(* Logix 5000 project; controller MV vendor 1 type 14 code 217 rev 31.11; software revision 31.00; part 17 of 53 *)
(* tags used below, declared in another part *)
   Alarm_Reset : BOOL;
   CheckTimeMask : INT;
   CLOCKsetvalues : DINT[7];
   CurrentTime : DateTime;
   CWD : CHECKWORD_FLAGS;
   Delphi_Does_Eng_Func : BOOL;
   MC_CLOCK_system_set : BOOL;
   MC_CP1 : PlantItem;   // CP1
   MC_data_file_value_to_move : DINT;
   MC_GBYV1 : PlantItem;   // GBYV1
   MC_N10 : INT[255];   // SETTINGS
   MC_N200 : INT[255];   // CHK_WORK Plant item fault che cking work area
   MC_N255 : INT[255];   // CHECKWORDS Plant item checkword s
   MC_P1 : PlantItem;   // P1
   MC_P2 : PlantItem;   // P2
   MC_P3 : PlantItem;   // P3
   MC_P4 : PlantItem;   // P4
   MC_SFile : INT[255];   // SLC Equivalent System File, So Original Code Can Remain
   MC_SP_R1_1 : PlantItem;   // SP_R1_1
   MC_SP_R2_1 : PlantItem;   // SP_R2_1
   MC_SP_R3_1 : PlantItem;   // SP_R3_1
   MC_T4 : TIMER[255];   // TIMER
   TempChecktime : DINT;
(* MC_Common, continued *)

ROUTINE MC_ITEMCHECK_200   (* ladder *)
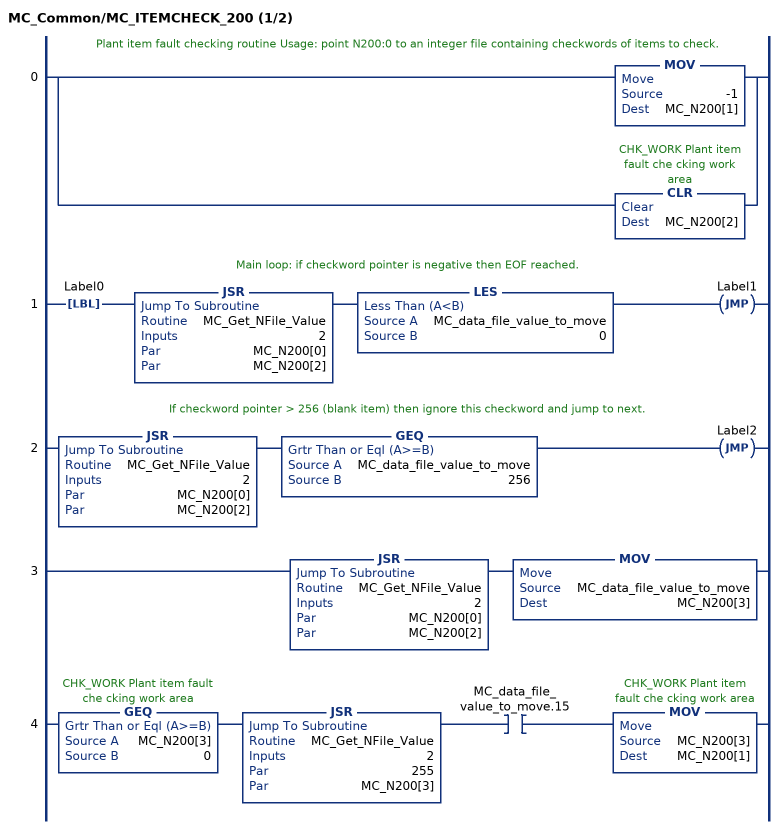
   // Plant item fault checking routine Usage: point N200:0 to an integer file containing checkwords of items to check.
   0: [MOV(-1,MC_N200[1]) ,CLR(MC_N200[2]) ];
   // Main loop: if checkword pointer is negative then EOF reached.
   1: LBL(Label0)JSR(MC_Get_NFile_Value,2,MC_N200[0],MC_N200[2])LES(MC_data_file_value_to_move,0)JMP(Label1);
   // If checkword pointer > 256 (blank item) then ignore this checkword and jump to next.
   2: JSR(MC_Get_NFile_Value,2,MC_N200[0],MC_N200[2])GEQ(MC_data_file_value_to_move,256)JMP(Label2);
   3: JSR(MC_Get_NFile_Value,2,MC_N200[0],MC_N200[2])MOV(MC_data_file_value_to_move,MC_N200[3]);
   4: GEQ(MC_N200[3],0)JSR(MC_Get_NFile_Value,2,255,MC_N200[3])XIC(MC_data_file_value_to_move.15)MOV(MC_N200[3],MC_N200[1]);
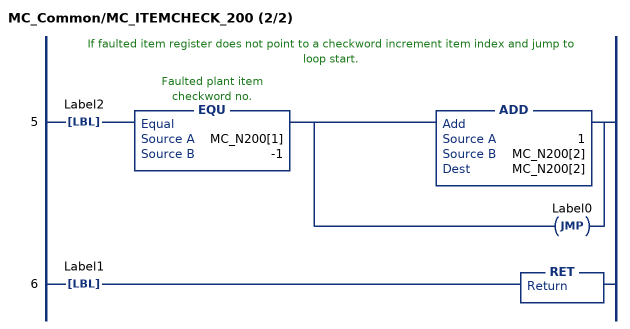
   // If faulted item register does not point to a checkword increment item index and jump to loop start.
   5: LBL(Label2)EQU(MC_N200[1],-1)[ADD(1,MC_N200[2],MC_N200[2]) ,JMP(Label0) ];
   6: LBL(Label1)RET();
END_ROUTINE

ROUTINE MC_MAIN   (* ladder *)
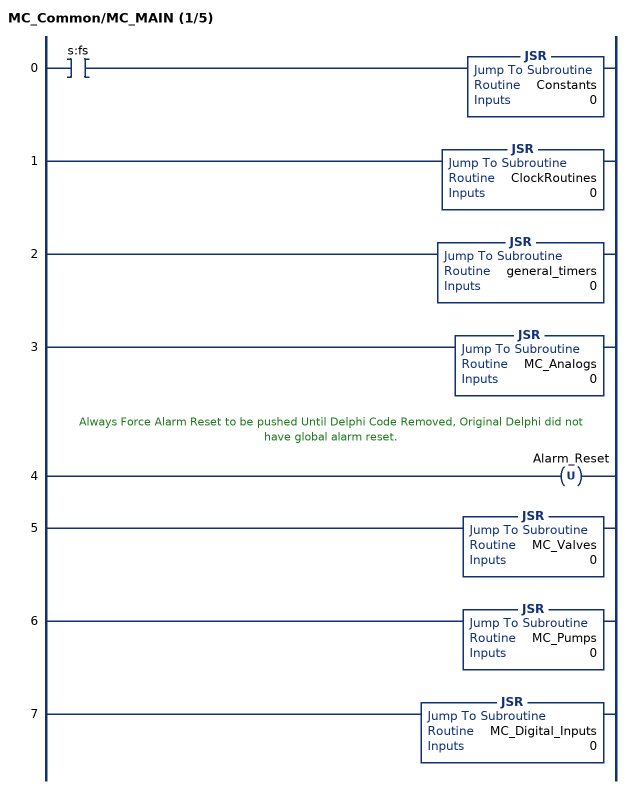
   0: XIC(s:fs)JSR(Constants,0);
   1: JSR(ClockRoutines,0);
   2: JSR(general_timers,0);
   3: JSR(MC_Analogs,0);
   // Always Force Alarm Reset to be pushed Until Delphi Code Removed, Original Delphi did not have global alarm reset.
   4: OTU(Alarm_Reset);
   5: JSR(MC_Valves,0);
   6: JSR(MC_Pumps,0);
   7: JSR(MC_Digital_Inputs,0);
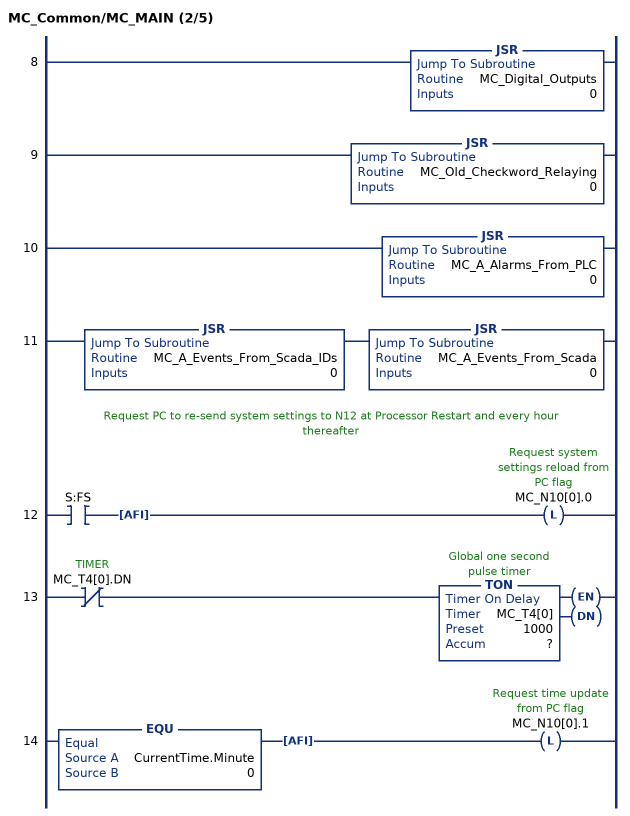
   8: JSR(MC_Digital_Outputs,0);
   9: JSR(MC_Old_Checkword_Relaying,0);
   10: JSR(MC_A_Alarms_From_PLC,0);
   11: JSR(MC_A_Events_From_Scada_IDs,0)JSR(MC_A_Events_From_Scada,0);
   // Request PC to re-send system settings to N12 at Processor Restart and every hour thereafter
   12: XIC(S:FS)AFI()OTL(MC_N10[0].0);
   13: XIO(MC_T4[0].DN)TON(MC_T4[0],?,?);
   14: EQU(CurrentTime.Minute,0)AFI()OTL(MC_N10[0].1);
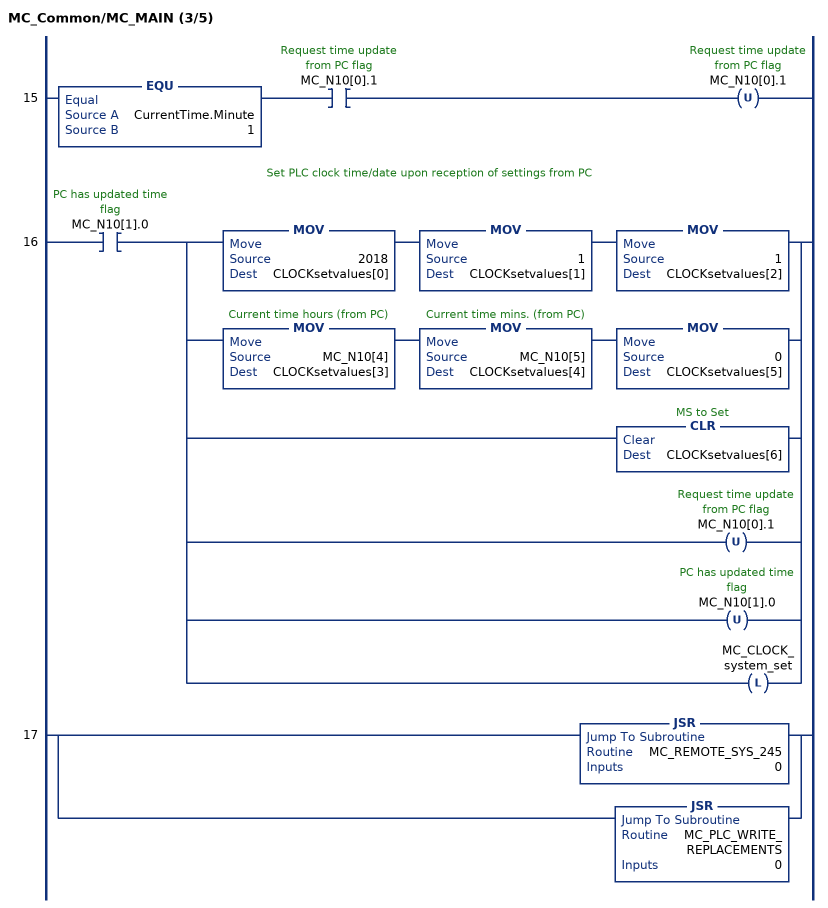
   15: EQU(CurrentTime.Minute,1)XIC(MC_N10[0].1)OTU(MC_N10[0].1);
   // Set PLC clock time/date upon reception of settings from PC
   16: XIC(MC_N10[1].0)[MOV(2018,CLOCKsetvalues[0]) MOV(1,CLOCKsetvalues[1]) MOV(1,CLOCKsetvalues[2]) ,MOV(MC_N10[4],CLOCKsetvalues[3]) MOV(MC_N10[5],CLOCKsetvalues[4]) MOV(0,CLOCKsetvalues[5]) ,CLR(CLOCKsetvalues[6]) ,OTU(MC_N10[0].1) ,OTU(MC_N10[1].0) ,OTL(MC_CLOCK_system_set) ];
   17: [JSR(MC_REMOTE_SYS_245,0) ,JSR(MC_PLC_WRITE_REPLACEMENTS,0) ];
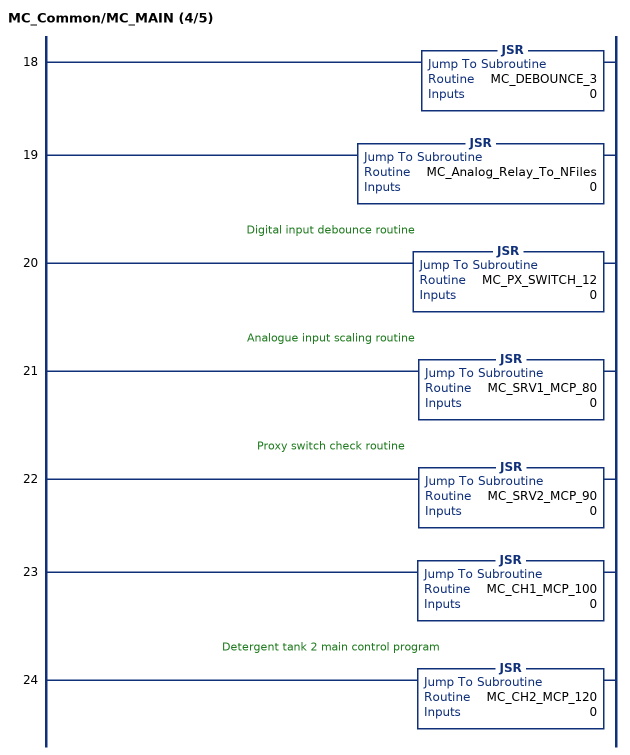
   18: JSR(MC_DEBOUNCE_3,0);
   19: JSR(MC_Analog_Relay_To_NFiles,0);
   // Digital input debounce routine
   20: JSR(MC_PX_SWITCH_12,0);
   // Analogue input scaling routine
   21: JSR(MC_SRV1_MCP_80,0);
   // Proxy switch check routine
   22: JSR(MC_SRV2_MCP_90,0);
   23: JSR(MC_CH1_MCP_100,0);
   // Detergent tank 2 main control program
   24: JSR(MC_CH2_MCP_120,0);
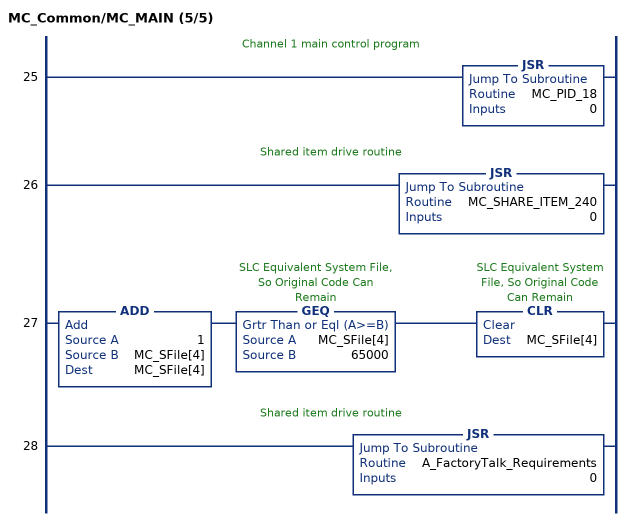
   // Channel 1 main control program
   25: JSR(MC_PID_18,0);
   // Shared item drive routine
   26: JSR(MC_SHARE_ITEM_240,0);
   27: ADD(1,MC_SFile[4],MC_SFile[4])GEQ(MC_SFile[4],65000)CLR(MC_SFile[4]);
   // Shared item drive routine
   28: JSR(A_FactoryTalk_Requirements,0);
END_ROUTINE

ROUTINE MC_Old_Checkword_Relaying   (* ladder *)
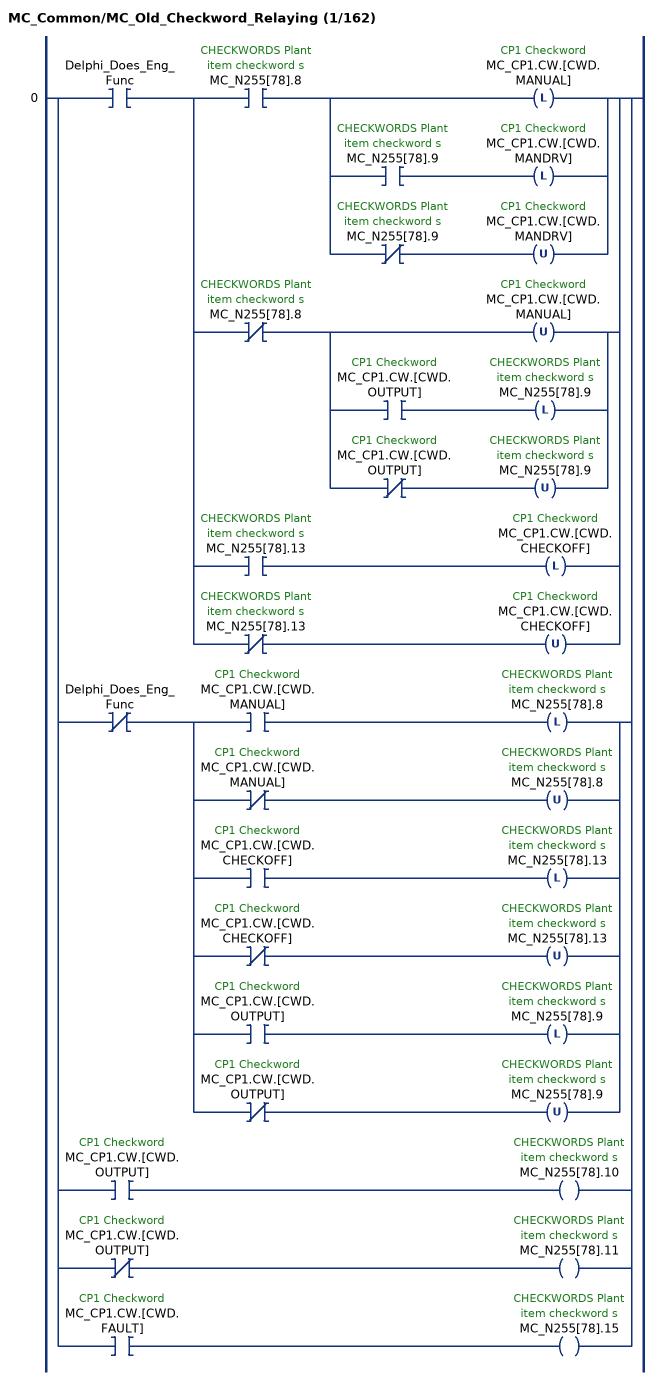
   0: [XIC(Delphi_Does_Eng_Func) [[XIC(MC_N255[78].8) [OTL(MC_CP1.CW.[CWD.MANUAL]) ,XIC(MC_N255[78].9) OTL(MC_CP1.CW.[CWD.MANDRV]) ,XIO(MC_N255[78].9) OTU(MC_CP1.CW.[CWD.MANDRV]) ] ,XIO(MC_N255[78].8) [OTU(MC_CP1.CW.[CWD.MANUAL]) ,[XIC(MC_CP1.CW.[CWD.OUTPUT]) OTL(MC_N255[78].9) ,XIO(MC_CP1.CW.[CWD.OUTPUT]) OTU(MC_N255[78].9) ] ] ] ,[XIC(MC_N255[78].13) OTL(MC_CP1.CW.[CWD.CHECKOFF]) ,XIO(MC_N255[78].13) OTU(MC_CP1.CW.[CWD.CHECKOFF]) ] ] ,XIO(Delphi_Does_Eng_Func) [[XIC(MC_CP1.CW.[CWD.MANUAL]) OTL(MC_N255[78].8) ,XIO(MC_CP1.CW.[CWD.MANUAL]) OTU(MC_N255[78].8) ] ,[XIC(MC_CP1.CW.[CWD.CHECKOFF]) OTL(MC_N255[78].13) ,XIO(MC_CP1.CW.[CWD.CHECKOFF]) OTU(MC_N255[78].13) ] ,[XIC(MC_CP1.CW.[CWD.OUTPUT]) OTL(MC_N255[78].9) ,XIO(MC_CP1.CW.[CWD.OUTPUT]) OTU(MC_N255[78].9) ] ] ,XIC(MC_CP1.CW.[CWD.OUTPUT]) OTE(MC_N255[78].10) ,XIO(MC_CP1.CW.[CWD.OUTPUT]) OTE(MC_N255[78].11) ,XIC(MC_CP1.CW.[CWD.FAULT]) OTE(MC_N255[78].15) ];
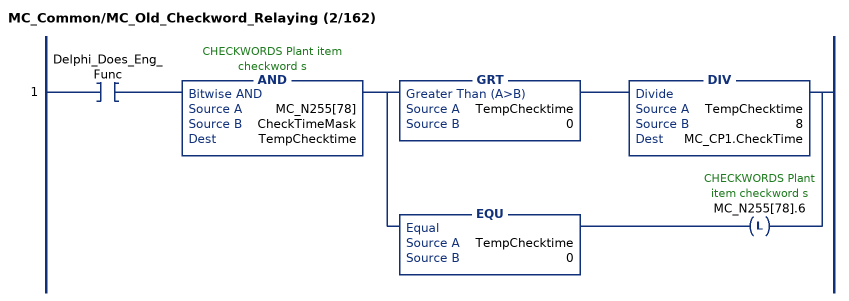
   1: XIC(Delphi_Does_Eng_Func)AND(MC_N255[78],CheckTimeMask,TempChecktime)[GRT(TempChecktime,0) DIV(TempChecktime,8,MC_CP1.CheckTime) ,EQU(TempChecktime,0) OTL(MC_N255[78].6) ];
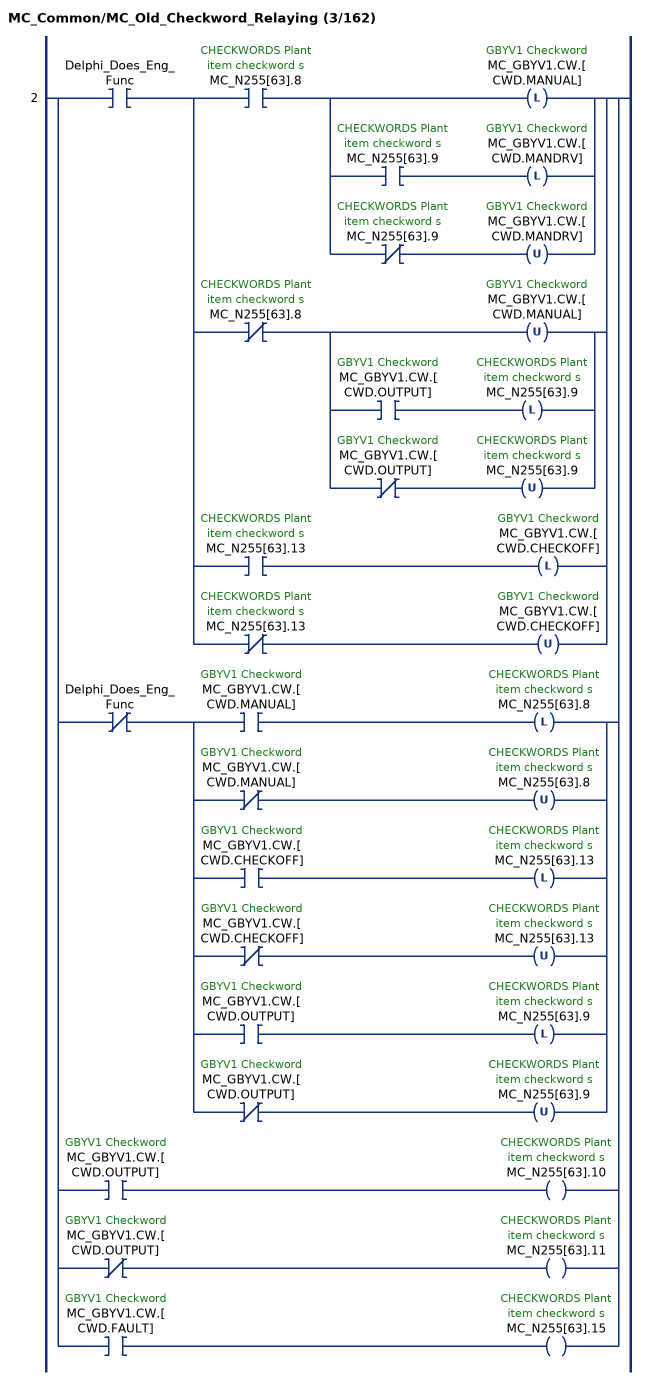
   2: [XIC(Delphi_Does_Eng_Func) [[XIC(MC_N255[63].8) [OTL(MC_GBYV1.CW.[CWD.MANUAL]) ,XIC(MC_N255[63].9) OTL(MC_GBYV1.CW.[CWD.MANDRV]) ,XIO(MC_N255[63].9) OTU(MC_GBYV1.CW.[CWD.MANDRV]) ] ,XIO(MC_N255[63].8) [OTU(MC_GBYV1.CW.[CWD.MANUAL]) ,[XIC(MC_GBYV1.CW.[CWD.OUTPUT]) OTL(MC_N255[63].9) ,XIO(MC_GBYV1.CW.[CWD.OUTPUT]) OTU(MC_N255[63].9) ] ] ] ,[XIC(MC_N255[63].13) OTL(MC_GBYV1.CW.[CWD.CHECKOFF]) ,XIO(MC_N255[63].13) OTU(MC_GBYV1.CW.[CWD.CHECKOFF]) ] ] ,XIO(Delphi_Does_Eng_Func) [[XIC(MC_GBYV1.CW.[CWD.MANUAL]) OTL(MC_N255[63].8) ,XIO(MC_GBYV1.CW.[CWD.MANUAL]) OTU(MC_N255[63].8) ] ,[XIC(MC_GBYV1.CW.[CWD.CHECKOFF]) OTL(MC_N255[63].13) ,XIO(MC_GBYV1.CW.[CWD.CHECKOFF]) OTU(MC_N255[63].13) ] ,[XIC(MC_GBYV1.CW.[CWD.OUTPUT]) OTL(MC_N255[63].9) ,XIO(MC_GBYV1.CW.[CWD.OUTPUT]) OTU(MC_N255[63].9) ] ] ,XIC(MC_GBYV1.CW.[CWD.OUTPUT]) OTE(MC_N255[63].10) ,XIO(MC_GBYV1.CW.[CWD.OUTPUT]) OTE(MC_N255[63].11) ,XIC(MC_GBYV1.CW.[CWD.FAULT]) OTE(MC_N255[63].15) ];
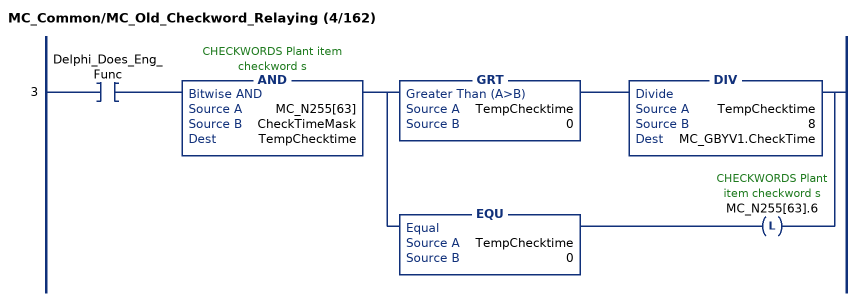
   3: XIC(Delphi_Does_Eng_Func)AND(MC_N255[63],CheckTimeMask,TempChecktime)[GRT(TempChecktime,0) DIV(TempChecktime,8,MC_GBYV1.CheckTime) ,EQU(TempChecktime,0) OTL(MC_N255[63].6) ];
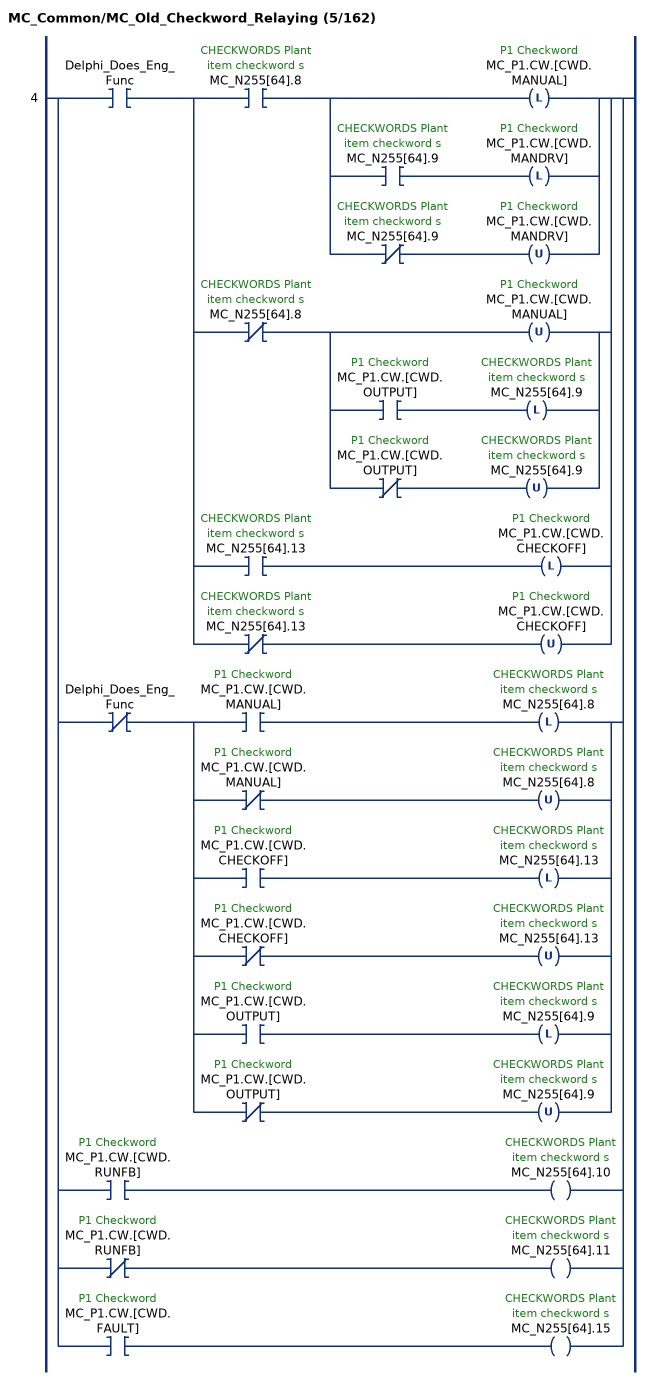
   4: [XIC(Delphi_Does_Eng_Func) [[XIC(MC_N255[64].8) [OTL(MC_P1.CW.[CWD.MANUAL]) ,XIC(MC_N255[64].9) OTL(MC_P1.CW.[CWD.MANDRV]) ,XIO(MC_N255[64].9) OTU(MC_P1.CW.[CWD.MANDRV]) ] ,XIO(MC_N255[64].8) [OTU(MC_P1.CW.[CWD.MANUAL]) ,[XIC(MC_P1.CW.[CWD.OUTPUT]) OTL(MC_N255[64].9) ,XIO(MC_P1.CW.[CWD.OUTPUT]) OTU(MC_N255[64].9) ] ] ] ,[XIC(MC_N255[64].13) OTL(MC_P1.CW.[CWD.CHECKOFF]) ,XIO(MC_N255[64].13) OTU(MC_P1.CW.[CWD.CHECKOFF]) ] ] ,XIO(Delphi_Does_Eng_Func) [[XIC(MC_P1.CW.[CWD.MANUAL]) OTL(MC_N255[64].8) ,XIO(MC_P1.CW.[CWD.MANUAL]) OTU(MC_N255[64].8) ] ,[XIC(MC_P1.CW.[CWD.CHECKOFF]) OTL(MC_N255[64].13) ,XIO(MC_P1.CW.[CWD.CHECKOFF]) OTU(MC_N255[64].13) ] ,[XIC(MC_P1.CW.[CWD.OUTPUT]) OTL(MC_N255[64].9) ,XIO(MC_P1.CW.[CWD.OUTPUT]) OTU(MC_N255[64].9) ] ] ,XIC(MC_P1.CW.[CWD.RUNFB]) OTE(MC_N255[64].10) ,XIO(MC_P1.CW.[CWD.RUNFB]) OTE(MC_N255[64].11) ,XIC(MC_P1.CW.[CWD.FAULT]) OTE(MC_N255[64].15) ];
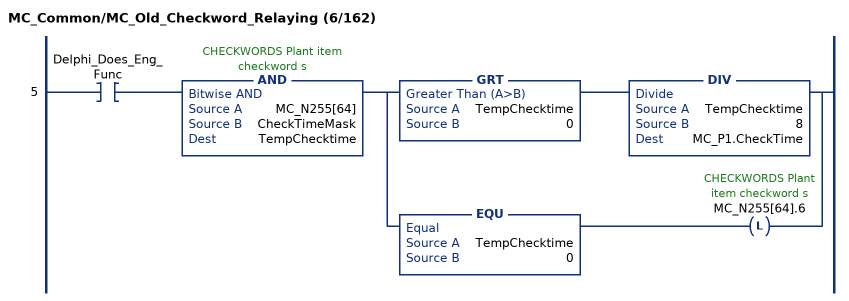
   5: XIC(Delphi_Does_Eng_Func)AND(MC_N255[64],CheckTimeMask,TempChecktime)[GRT(TempChecktime,0) DIV(TempChecktime,8,MC_P1.CheckTime) ,EQU(TempChecktime,0) OTL(MC_N255[64].6) ];
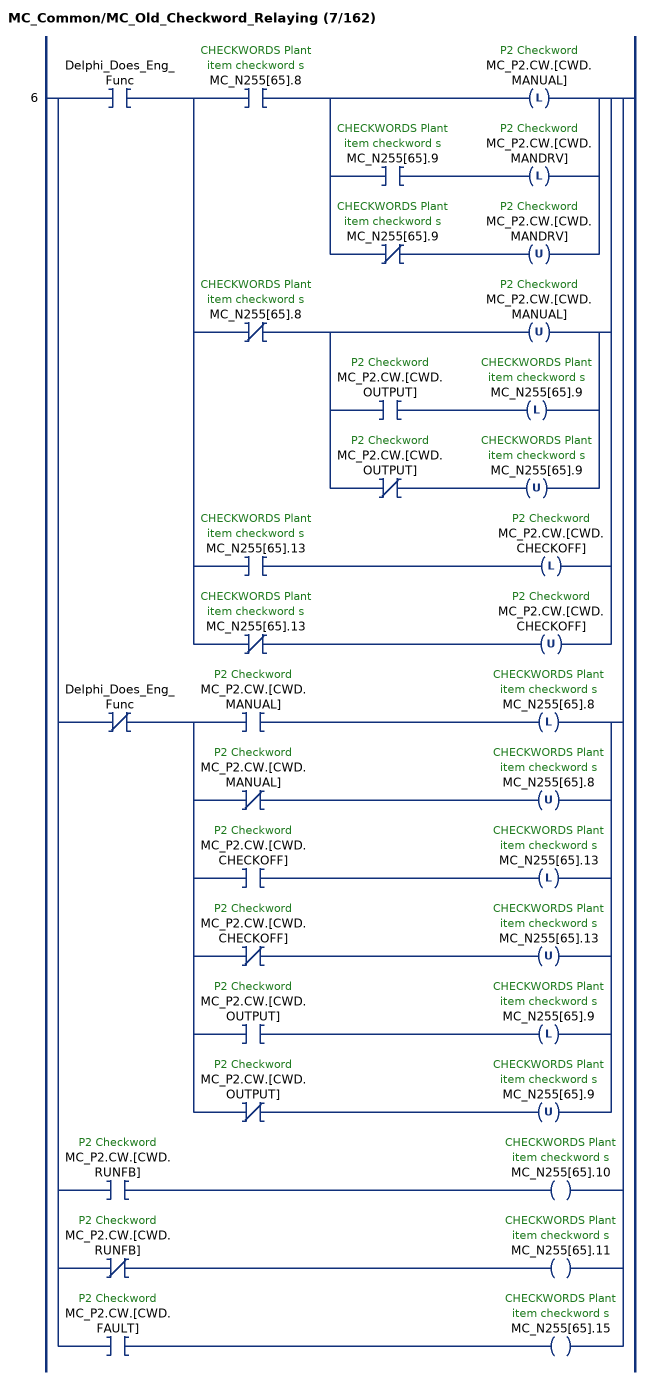
   6: [XIC(Delphi_Does_Eng_Func) [[XIC(MC_N255[65].8) [OTL(MC_P2.CW.[CWD.MANUAL]) ,XIC(MC_N255[65].9) OTL(MC_P2.CW.[CWD.MANDRV]) ,XIO(MC_N255[65].9) OTU(MC_P2.CW.[CWD.MANDRV]) ] ,XIO(MC_N255[65].8) [OTU(MC_P2.CW.[CWD.MANUAL]) ,[XIC(MC_P2.CW.[CWD.OUTPUT]) OTL(MC_N255[65].9) ,XIO(MC_P2.CW.[CWD.OUTPUT]) OTU(MC_N255[65].9) ] ] ] ,[XIC(MC_N255[65].13) OTL(MC_P2.CW.[CWD.CHECKOFF]) ,XIO(MC_N255[65].13) OTU(MC_P2.CW.[CWD.CHECKOFF]) ] ] ,XIO(Delphi_Does_Eng_Func) [[XIC(MC_P2.CW.[CWD.MANUAL]) OTL(MC_N255[65].8) ,XIO(MC_P2.CW.[CWD.MANUAL]) OTU(MC_N255[65].8) ] ,[XIC(MC_P2.CW.[CWD.CHECKOFF]) OTL(MC_N255[65].13) ,XIO(MC_P2.CW.[CWD.CHECKOFF]) OTU(MC_N255[65].13) ] ,[XIC(MC_P2.CW.[CWD.OUTPUT]) OTL(MC_N255[65].9) ,XIO(MC_P2.CW.[CWD.OUTPUT]) OTU(MC_N255[65].9) ] ] ,XIC(MC_P2.CW.[CWD.RUNFB]) OTE(MC_N255[65].10) ,XIO(MC_P2.CW.[CWD.RUNFB]) OTE(MC_N255[65].11) ,XIC(MC_P2.CW.[CWD.FAULT]) OTE(MC_N255[65].15) ];
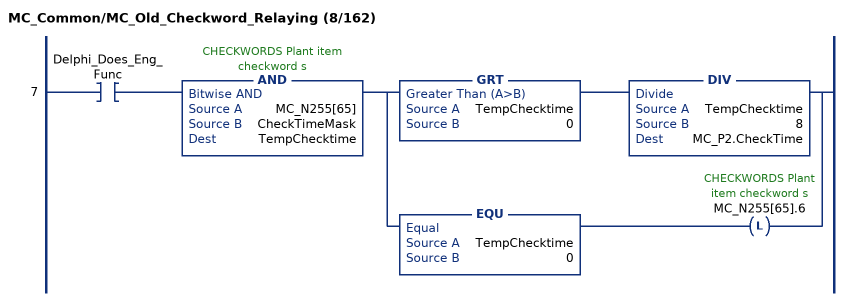
   7: XIC(Delphi_Does_Eng_Func)AND(MC_N255[65],CheckTimeMask,TempChecktime)[GRT(TempChecktime,0) DIV(TempChecktime,8,MC_P2.CheckTime) ,EQU(TempChecktime,0) OTL(MC_N255[65].6) ];
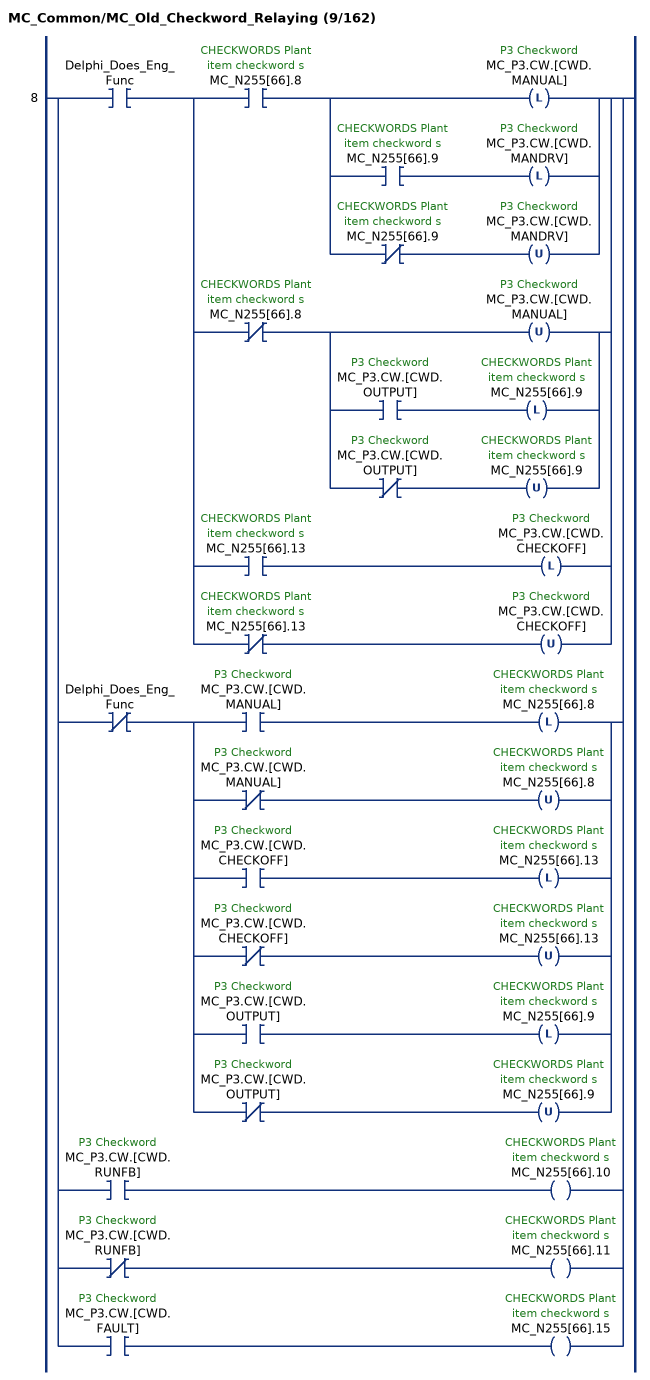
   8: [XIC(Delphi_Does_Eng_Func) [[XIC(MC_N255[66].8) [OTL(MC_P3.CW.[CWD.MANUAL]) ,XIC(MC_N255[66].9) OTL(MC_P3.CW.[CWD.MANDRV]) ,XIO(MC_N255[66].9) OTU(MC_P3.CW.[CWD.MANDRV]) ] ,XIO(MC_N255[66].8) [OTU(MC_P3.CW.[CWD.MANUAL]) ,[XIC(MC_P3.CW.[CWD.OUTPUT]) OTL(MC_N255[66].9) ,XIO(MC_P3.CW.[CWD.OUTPUT]) OTU(MC_N255[66].9) ] ] ] ,[XIC(MC_N255[66].13) OTL(MC_P3.CW.[CWD.CHECKOFF]) ,XIO(MC_N255[66].13) OTU(MC_P3.CW.[CWD.CHECKOFF]) ] ] ,XIO(Delphi_Does_Eng_Func) [[XIC(MC_P3.CW.[CWD.MANUAL]) OTL(MC_N255[66].8) ,XIO(MC_P3.CW.[CWD.MANUAL]) OTU(MC_N255[66].8) ] ,[XIC(MC_P3.CW.[CWD.CHECKOFF]) OTL(MC_N255[66].13) ,XIO(MC_P3.CW.[CWD.CHECKOFF]) OTU(MC_N255[66].13) ] ,[XIC(MC_P3.CW.[CWD.OUTPUT]) OTL(MC_N255[66].9) ,XIO(MC_P3.CW.[CWD.OUTPUT]) OTU(MC_N255[66].9) ] ] ,XIC(MC_P3.CW.[CWD.RUNFB]) OTE(MC_N255[66].10) ,XIO(MC_P3.CW.[CWD.RUNFB]) OTE(MC_N255[66].11) ,XIC(MC_P3.CW.[CWD.FAULT]) OTE(MC_N255[66].15) ];
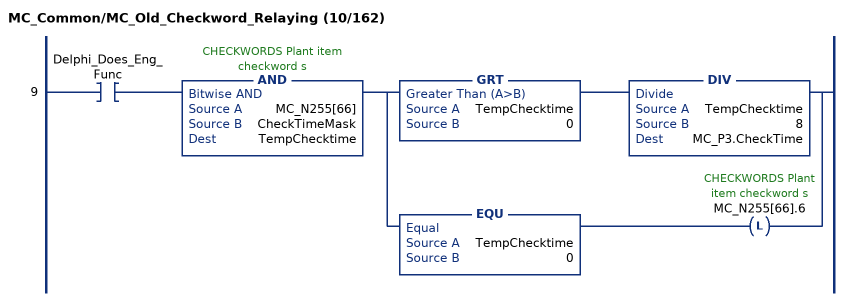
   9: XIC(Delphi_Does_Eng_Func)AND(MC_N255[66],CheckTimeMask,TempChecktime)[GRT(TempChecktime,0) DIV(TempChecktime,8,MC_P3.CheckTime) ,EQU(TempChecktime,0) OTL(MC_N255[66].6) ];
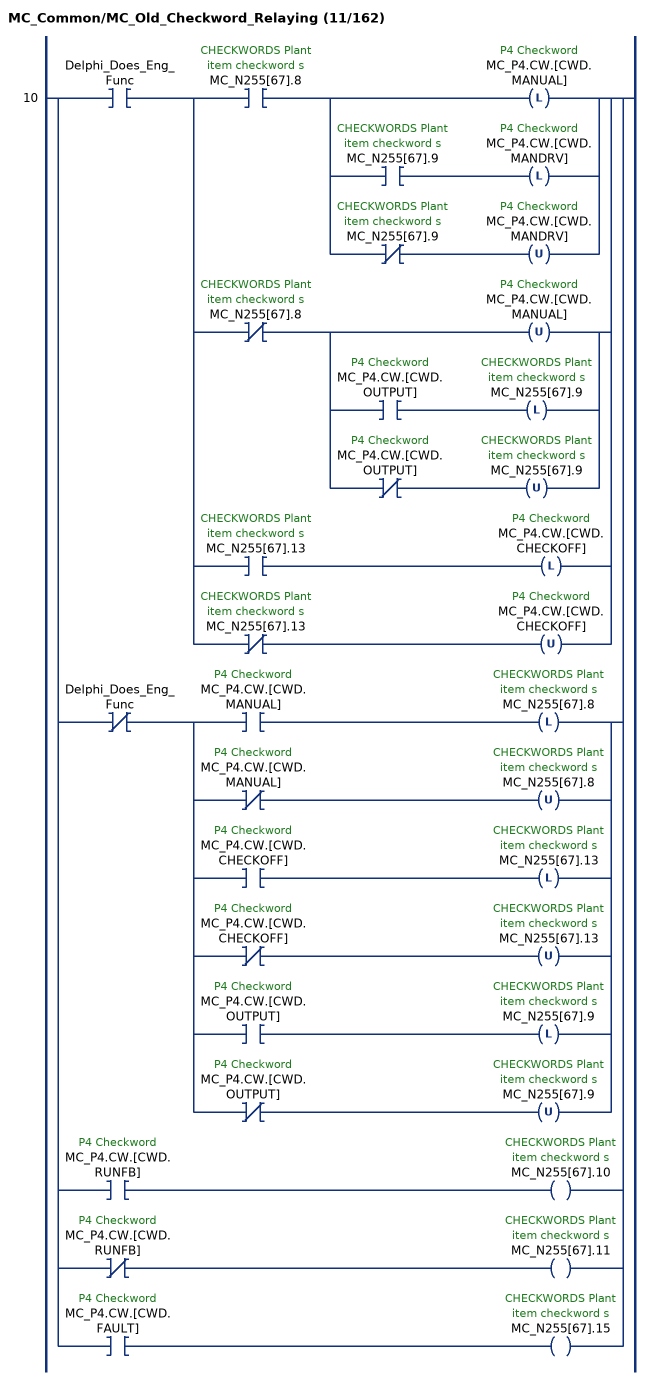
   10: [XIC(Delphi_Does_Eng_Func) [[XIC(MC_N255[67].8) [OTL(MC_P4.CW.[CWD.MANUAL]) ,XIC(MC_N255[67].9) OTL(MC_P4.CW.[CWD.MANDRV]) ,XIO(MC_N255[67].9) OTU(MC_P4.CW.[CWD.MANDRV]) ] ,XIO(MC_N255[67].8) [OTU(MC_P4.CW.[CWD.MANUAL]) ,[XIC(MC_P4.CW.[CWD.OUTPUT]) OTL(MC_N255[67].9) ,XIO(MC_P4.CW.[CWD.OUTPUT]) OTU(MC_N255[67].9) ] ] ] ,[XIC(MC_N255[67].13) OTL(MC_P4.CW.[CWD.CHECKOFF]) ,XIO(MC_N255[67].13) OTU(MC_P4.CW.[CWD.CHECKOFF]) ] ] ,XIO(Delphi_Does_Eng_Func) [[XIC(MC_P4.CW.[CWD.MANUAL]) OTL(MC_N255[67].8) ,XIO(MC_P4.CW.[CWD.MANUAL]) OTU(MC_N255[67].8) ] ,[XIC(MC_P4.CW.[CWD.CHECKOFF]) OTL(MC_N255[67].13) ,XIO(MC_P4.CW.[CWD.CHECKOFF]) OTU(MC_N255[67].13) ] ,[XIC(MC_P4.CW.[CWD.OUTPUT]) OTL(MC_N255[67].9) ,XIO(MC_P4.CW.[CWD.OUTPUT]) OTU(MC_N255[67].9) ] ] ,XIC(MC_P4.CW.[CWD.RUNFB]) OTE(MC_N255[67].10) ,XIO(MC_P4.CW.[CWD.RUNFB]) OTE(MC_N255[67].11) ,XIC(MC_P4.CW.[CWD.FAULT]) OTE(MC_N255[67].15) ];
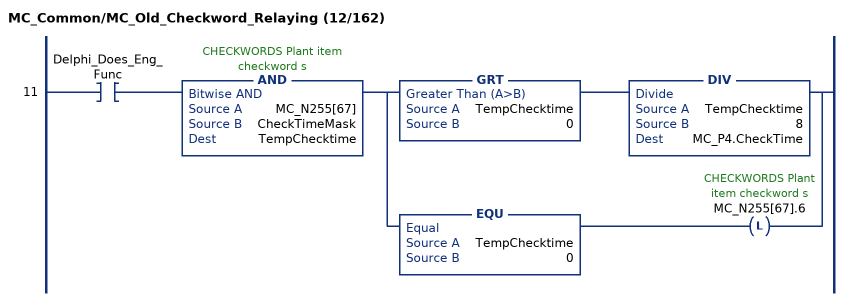
   11: XIC(Delphi_Does_Eng_Func)AND(MC_N255[67],CheckTimeMask,TempChecktime)[GRT(TempChecktime,0) DIV(TempChecktime,8,MC_P4.CheckTime) ,EQU(TempChecktime,0) OTL(MC_N255[67].6) ];
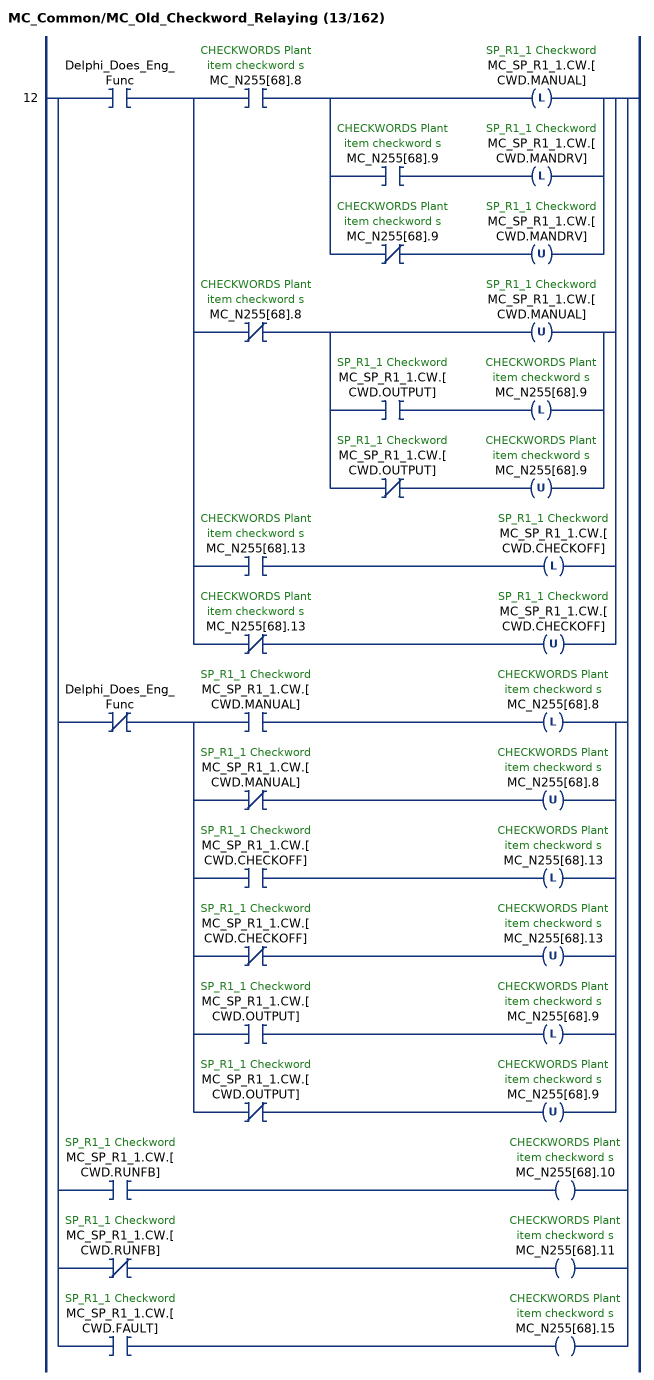
   12: [XIC(Delphi_Does_Eng_Func) [[XIC(MC_N255[68].8) [OTL(MC_SP_R1_1.CW.[CWD.MANUAL]) ,XIC(MC_N255[68].9) OTL(MC_SP_R1_1.CW.[CWD.MANDRV]) ,XIO(MC_N255[68].9) OTU(MC_SP_R1_1.CW.[CWD.MANDRV]) ] ,XIO(MC_N255[68].8) [OTU(MC_SP_R1_1.CW.[CWD.MANUAL]) ,[XIC(MC_SP_R1_1.CW.[CWD.OUTPUT]) OTL(MC_N255[68].9) ,XIO(MC_SP_R1_1.CW.[CWD.OUTPUT]) OTU(MC_N255[68].9) ] ] ] ,[XIC(MC_N255[68].13) OTL(MC_SP_R1_1.CW.[CWD.CHECKOFF]) ,XIO(MC_N255[68].13) OTU(MC_SP_R1_1.CW.[CWD.CHECKOFF]) ] ] ,XIO(Delphi_Does_Eng_Func) [[XIC(MC_SP_R1_1.CW.[CWD.MANUAL]) OTL(MC_N255[68].8) ,XIO(MC_SP_R1_1.CW.[CWD.MANUAL]) OTU(MC_N255[68].8) ] ,[XIC(MC_SP_R1_1.CW.[CWD.CHECKOFF]) OTL(MC_N255[68].13) ,XIO(MC_SP_R1_1.CW.[CWD.CHECKOFF]) OTU(MC_N255[68].13) ] ,[XIC(MC_SP_R1_1.CW.[CWD.OUTPUT]) OTL(MC_N255[68].9) ,XIO(MC_SP_R1_1.CW.[CWD.OUTPUT]) OTU(MC_N255[68].9) ] ] ,XIC(MC_SP_R1_1.CW.[CWD.RUNFB]) OTE(MC_N255[68].10) ,XIO(MC_SP_R1_1.CW.[CWD.RUNFB]) OTE(MC_N255[68].11) ,XIC(MC_SP_R1_1.CW.[CWD.FAULT]) OTE(MC_N255[68].15) ];
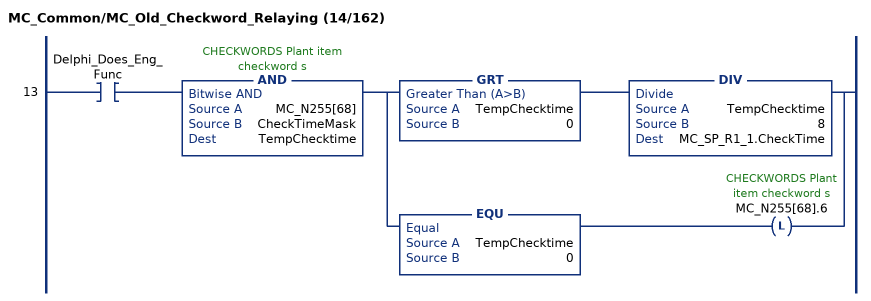
   13: XIC(Delphi_Does_Eng_Func)AND(MC_N255[68],CheckTimeMask,TempChecktime)[GRT(TempChecktime,0) DIV(TempChecktime,8,MC_SP_R1_1.CheckTime) ,EQU(TempChecktime,0) OTL(MC_N255[68].6) ];
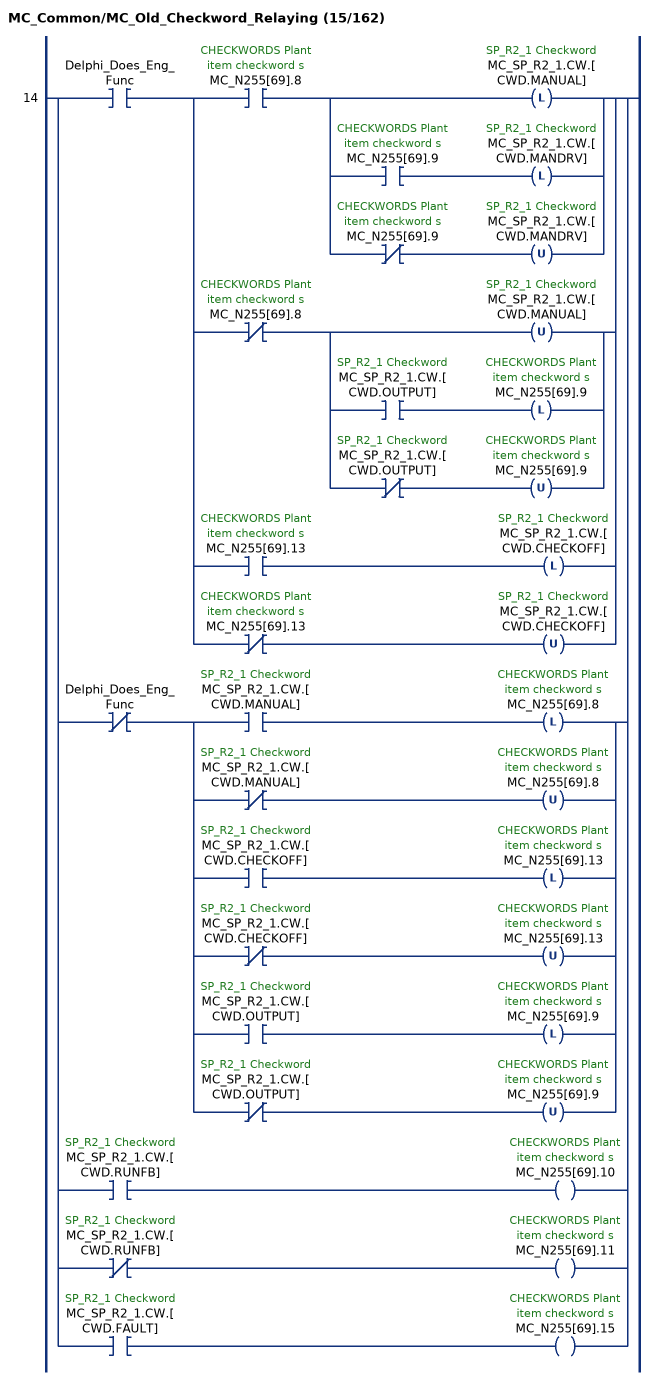
   14: [XIC(Delphi_Does_Eng_Func) [[XIC(MC_N255[69].8) [OTL(MC_SP_R2_1.CW.[CWD.MANUAL]) ,XIC(MC_N255[69].9) OTL(MC_SP_R2_1.CW.[CWD.MANDRV]) ,XIO(MC_N255[69].9) OTU(MC_SP_R2_1.CW.[CWD.MANDRV]) ] ,XIO(MC_N255[69].8) [OTU(MC_SP_R2_1.CW.[CWD.MANUAL]) ,[XIC(MC_SP_R2_1.CW.[CWD.OUTPUT]) OTL(MC_N255[69].9) ,XIO(MC_SP_R2_1.CW.[CWD.OUTPUT]) OTU(MC_N255[69].9) ] ] ] ,[XIC(MC_N255[69].13) OTL(MC_SP_R2_1.CW.[CWD.CHECKOFF]) ,XIO(MC_N255[69].13) OTU(MC_SP_R2_1.CW.[CWD.CHECKOFF]) ] ] ,XIO(Delphi_Does_Eng_Func) [[XIC(MC_SP_R2_1.CW.[CWD.MANUAL]) OTL(MC_N255[69].8) ,XIO(MC_SP_R2_1.CW.[CWD.MANUAL]) OTU(MC_N255[69].8) ] ,[XIC(MC_SP_R2_1.CW.[CWD.CHECKOFF]) OTL(MC_N255[69].13) ,XIO(MC_SP_R2_1.CW.[CWD.CHECKOFF]) OTU(MC_N255[69].13) ] ,[XIC(MC_SP_R2_1.CW.[CWD.OUTPUT]) OTL(MC_N255[69].9) ,XIO(MC_SP_R2_1.CW.[CWD.OUTPUT]) OTU(MC_N255[69].9) ] ] ,XIC(MC_SP_R2_1.CW.[CWD.RUNFB]) OTE(MC_N255[69].10) ,XIO(MC_SP_R2_1.CW.[CWD.RUNFB]) OTE(MC_N255[69].11) ,XIC(MC_SP_R2_1.CW.[CWD.FAULT]) OTE(MC_N255[69].15) ];
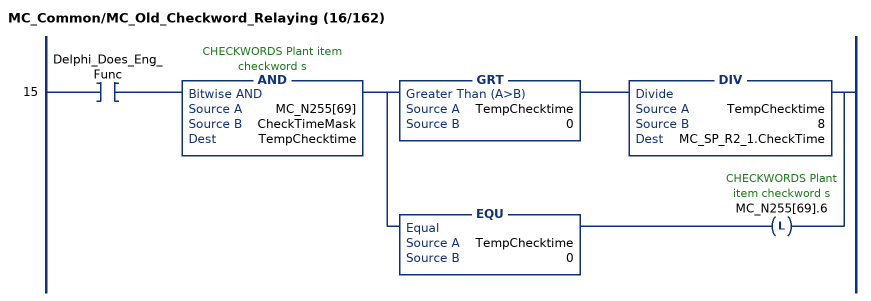
   15: XIC(Delphi_Does_Eng_Func)AND(MC_N255[69],CheckTimeMask,TempChecktime)[GRT(TempChecktime,0) DIV(TempChecktime,8,MC_SP_R2_1.CheckTime) ,EQU(TempChecktime,0) OTL(MC_N255[69].6) ];
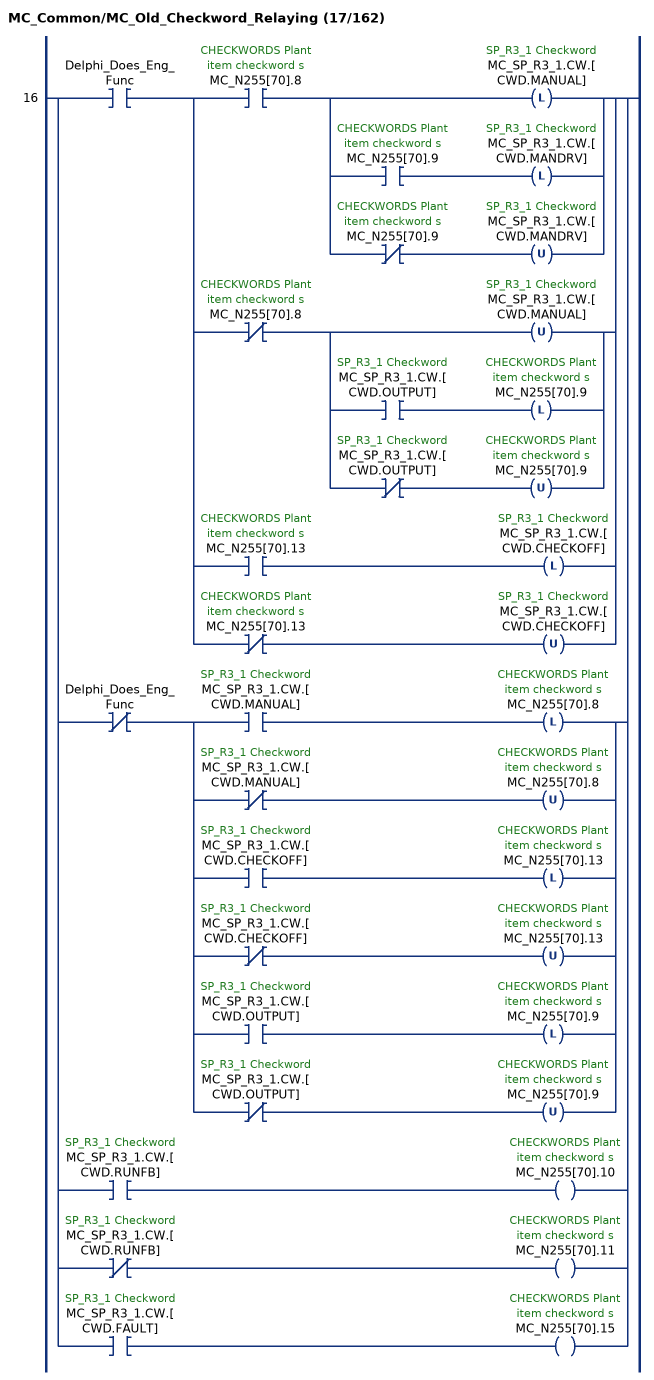
   16: [XIC(Delphi_Does_Eng_Func) [[XIC(MC_N255[70].8) [OTL(MC_SP_R3_1.CW.[CWD.MANUAL]) ,XIC(MC_N255[70].9) OTL(MC_SP_R3_1.CW.[CWD.MANDRV]) ,XIO(MC_N255[70].9) OTU(MC_SP_R3_1.CW.[CWD.MANDRV]) ] ,XIO(MC_N255[70].8) [OTU(MC_SP_R3_1.CW.[CWD.MANUAL]) ,[XIC(MC_SP_R3_1.CW.[CWD.OUTPUT]) OTL(MC_N255[70].9) ,XIO(MC_SP_R3_1.CW.[CWD.OUTPUT]) OTU(MC_N255[70].9) ] ] ] ,[XIC(MC_N255[70].13) OTL(MC_SP_R3_1.CW.[CWD.CHECKOFF]) ,XIO(MC_N255[70].13) OTU(MC_SP_R3_1.CW.[CWD.CHECKOFF]) ] ] ,XIO(Delphi_Does_Eng_Func) [[XIC(MC_SP_R3_1.CW.[CWD.MANUAL]) OTL(MC_N255[70].8) ,XIO(MC_SP_R3_1.CW.[CWD.MANUAL]) OTU(MC_N255[70].8) ] ,[XIC(MC_SP_R3_1.CW.[CWD.CHECKOFF]) OTL(MC_N255[70].13) ,XIO(MC_SP_R3_1.CW.[CWD.CHECKOFF]) OTU(MC_N255[70].13) ] ,[XIC(MC_SP_R3_1.CW.[CWD.OUTPUT]) OTL(MC_N255[70].9) ,XIO(MC_SP_R3_1.CW.[CWD.OUTPUT]) OTU(MC_N255[70].9) ] ] ,XIC(MC_SP_R3_1.CW.[CWD.RUNFB]) OTE(MC_N255[70].10) ,XIO(MC_SP_R3_1.CW.[CWD.RUNFB]) OTE(MC_N255[70].11) ,XIC(MC_SP_R3_1.CW.[CWD.FAULT]) OTE(MC_N255[70].15) ];
